   3225: 'Carrier 50 Drive: PROFINET Setpoint timeout', class No Acknowledgement, trigger "DB302_HMI_Faults_Carrier50_Faults_1" bit 8
   3226: 'Carrier 50 Power unit: Overcurrent', class No Acknowledgement, trigger "DB302_HMI_Faults_Carrier50_Faults_1" bit 9
   3227: 'Carrier 50 Power unit: DC link voltage overvoltage', class No Acknowledgement, trigger "DB302_HMI_Faults_Carrier50_Faults_1" bit 10
   3228: 'Carrier 50 Power unit: DC link voltage undervoltage', class No Acknowledgement, trigger "DB302_HMI_Faults_Carrier50_Faults_1" bit 11
   3229: 'Carrier 50 Power unit: Line phase failure in main circuit', class No Acknowledgement, trigger "DB302_HMI_Faults_Carrier50_Faults_1" bit 12
   3230: 'Carrier 50 Power unit: Phase failure motor cable', class No Acknowledgement, trigger "DB302_HMI_Faults_Carrier50_Faults_1" bit 13
   3231: 'Carrier 50 Power unit: Ground fault', class No Acknowledgement, trigger "DB302_HMI_Faults_Carrier50_Faults_1" bit 14
   3232: 'Spare_Fault_3232', class No Acknowledgement, trigger "DB302_HMI_Faults_Carrier50_Faults_1" bit 15
   3233: 'Carrier 50 Motion Off Fault', class No Acknowledgement, trigger "DB302_HMI_Faults_Carrier50_Faults_2" bit 0
   3234: 'Carrier 50 Motion On Fault', class No Acknowledgement, trigger "DB302_HMI_Faults_Carrier50_Faults_2" bit 1
   3235: 'Carrier 50 Spacing Fault', class No Acknowledgement, trigger "DB302_HMI_Faults_Carrier50_Faults_2" bit 2
   3236: 'Carrier 50 Duplicate Carrier Number Fault', class No Acknowledgement, trigger "DB302_HMI_Faults_Carrier50_Faults_2" bit 3
   3237: 'Spare_Fault_3237', class No Acknowledgement, trigger "DB302_HMI_Faults_Carrier50_Faults_2" bit 4
   3238: 'Spare_Fault_3238', class No Acknowledgement, trigger "DB302_HMI_Faults_Carrier50_Faults_2" bit 5
   3239: 'Spare_Fault_3239', class No Acknowledgement, trigger "DB302_HMI_Faults_Carrier50_Faults_2" bit 6
   3240: 'Spare_Fault_3240', class No Acknowledgement, trigger "DB302_HMI_Faults_Carrier50_Faults_2" bit 7
   3241: 'Spare_Fault_3241', class No Acknowledgement, trigger "DB302_HMI_Faults_Carrier50_Faults_2" bit 8
   3242: 'Spare_Fault_3242', class No Acknowledgement, trigger "DB302_HMI_Faults_Carrier50_Faults_2" bit 9
   3243: 'Spare_Fault_3243', class No Acknowledgement, trigger "DB302_HMI_Faults_Carrier50_Faults_2" bit 10
   3244: 'Spare_Fault_3244', class No Acknowledgement, trigger "DB302_HMI_Faults_Carrier50_Faults_2" bit 11
   3245: 'Spare_Fault_3245', class No Acknowledgement, trigger "DB302_HMI_Faults_Carrier50_Faults_2" bit 12
   3246: 'Spare_Fault_3246', class No Acknowledgement, trigger "DB302_HMI_Faults_Carrier50_Faults_2" bit 13
   3247: 'Spare_Fault_3247', class No Acknowledgement, trigger "DB302_HMI_Faults_Carrier50_Faults_2" bit 14
   3248: 'Spare_Fault_3248', class No Acknowledgement, trigger "DB302_HMI_Faults_Carrier50_Faults_2" bit 15
   3249: 'Spare_Fault_3249', class No Acknowledgement, trigger "DB302_HMI_Faults_Carrier50_Faults_3" bit 0
   3250: 'Spare_Fault_3250', class No Acknowledgement, trigger "DB302_HMI_Faults_Carrier50_Faults_3" bit 1
   3251: 'Spare_Fault_3251', class No Acknowledgement, trigger "DB302_HMI_Faults_Carrier50_Faults_3" bit 2
   3252: 'Spare_Fault_3252', class No Acknowledgement, trigger "DB302_HMI_Faults_Carrier50_Faults_3" bit 3
   3253: 'Spare_Fault_3253', class No Acknowledgement, trigger "DB302_HMI_Faults_Carrier50_Faults_3" bit 4
   3254: 'Spare_Fault_3254', class No Acknowledgement, trigger "DB302_HMI_Faults_Carrier50_Faults_3" bit 5
   3255: 'Spare_Fault_3255', class No Acknowledgement, trigger "DB302_HMI_Faults_Carrier50_Faults_3" bit 6
   3256: 'Spare_Fault_3256', class No Acknowledgement, trigger "DB302_HMI_Faults_Carrier50_Faults_3" bit 7
   3257: 'Spare_Fault_3257', class No Acknowledgement, trigger "DB302_HMI_Faults_Carrier50_Faults_3" bit 8
   3258: 'Spare_Fault_3258', class No Acknowledgement, trigger "DB302_HMI_Faults_Carrier50_Faults_3" bit 9
   3259: 'Spare_Fault_3259', class No Acknowledgement, trigger "DB302_HMI_Faults_Carrier50_Faults_3" bit 10
   3260: 'Spare_Fault_3260', class No Acknowledgement, trigger "DB302_HMI_Faults_Carrier50_Faults_3" bit 11
   3261: 'Spare_Fault_3261', class No Acknowledgement, trigger "DB302_HMI_Faults_Carrier50_Faults_3" bit 12
   3262: 'Spare_Fault_3262', class No Acknowledgement, trigger "DB302_HMI_Faults_Carrier50_Faults_3" bit 13
   3263: 'Spare_Fault_3263', class No Acknowledgement, trigger "DB302_HMI_Faults_Carrier50_Faults_3" bit 14
   3264: 'Spare_Fault_3264', class No Acknowledgement, trigger "DB302_HMI_Faults_Carrier50_Faults_3" bit 15
   3265: 'Carrier 51 Disconnect Open Power Fault DI11.0', class No Acknowledgement, trigger "DB302_HMI_Faults_Carrier51_Faults_0" bit 0
   3266: 'Carrier 51 Drive Profinet Comm Fault', class No Acknowledgement, trigger "DB302_HMI_Faults_Carrier51_Faults_0" bit 1
   3267: 'Carrier 51 Production Stop Not Reset', class No Acknowledgement, trigger "DB302_HMI_Faults_Carrier51_Faults_0" bit 2
   3268: 'Carrier 51 CB02122 Tripped', class No Acknowledgement, trigger "DB302_HMI_Faults_Carrier51_Faults_0" bit 3
   3269: 'Carrier 51 CB02123 Tripped', class No Acknowledgement, trigger "DB302_HMI_Faults_Carrier51_Faults_0" bit 4
   3270: 'Carrier 51 AUX1 CB Tripped', class No Acknowledgement, trigger "DB302_HMI_Faults_Carrier51_Faults_0" bit 5
   3271: 'Carrier 51 AUX2 CB Tripped', class No Acknowledgement, trigger "DB302_HMI_Faults_Carrier51_Faults_0" bit 6
   3272: 'Carrier 51 PLC Not Communicating', class No Acknowledgement, trigger "DB302_HMI_Faults_Carrier51_Faults_0" bit 7
   3273: 'Carrier 51 Safe Input Card Fault', class No Acknowledgement, trigger "DB302_HMI_Faults_Carrier51_Faults_0" bit 8
   3274: 'Carrier 51 Safe Output Card Fault', class No Acknowledgement, trigger "DB302_HMI_Faults_Carrier51_Faults_0" bit 9
   3275: 'Carrier 51 Standard Input Card Fault', class No Acknowledgement, trigger "DB302_HMI_Faults_Carrier51_Faults_0" bit 10
   3276: 'Carrier 51 Standard Output Card Fault', class No Acknowledgement, trigger "DB302_HMI_Faults_Carrier51_Faults_0" bit 11
   3277: 'Carrier 51 Encoder Position Fault', class No Acknowledgement, trigger "DB302_HMI_Faults_Carrier51_Faults_0" bit 12
   3278: 'Carrier 51 Encoder Internal Error', class No Acknowledgement, trigger "DB302_HMI_Faults_Carrier51_Faults_0" bit 13
   3279: 'Carrier 51 Encoder Comm Fault', class No Acknowledgement, trigger "DB302_HMI_Faults_Carrier51_Faults_0" bit 14
   3280: 'Carrier 51 HMI Comm Fault', class No Acknowledgement, trigger "DB302_HMI_Faults_Carrier51_Faults_0" bit 15
   3281: 'Carrier 51 Crash Detection Fault', class No Acknowledgement, trigger "DB302_HMI_Faults_Carrier51_Faults_1" bit 0
   3282: 'Carrier 51 Carrier Number Invalid', class No Acknowledgement, trigger "DB302_HMI_Faults_Carrier51_Faults_1" bit 1
   3283: 'Carrier 51 Drive: PROFINET configuration error', class No Acknowledgement, trigger "DB302_HMI_Faults_Carrier51_Faults_1" bit 2
   3284: 'Carrier 51 Drive: Error internal communications', class No Acknowledgement, trigger "DB302_HMI_Faults_Carrier51_Faults_1" bit 3
   3285: 'Carrier 51 Drive: Motor overtemperature', class No Acknowledgement, trigger "DB302_HMI_Faults_Carrier51_Faults_1" bit 4
   3286: 'Carrier 51 Drive: Motor overcurrent', class No Acknowledgement, trigger "DB302_HMI_Faults_Carrier51_Faults_1" bit 5
   3287: 'Carrier 51 Drive: Infeed or power unit not ready', class No Acknowledgement, trigger "DB302_HMI_Faults_Carrier51_Faults_1" bit 6
   3288: 'Carrier 51 Drive: Short-circuit/ground fault detected', class No Acknowledgement, trigger "DB302_HMI_Faults_Carrier51_Faults_1" bit 7
   3289: 'Carrier 51 Drive: PROFINET Setpoint timeout', class No Acknowledgement, trigger "DB302_HMI_Faults_Carrier51_Faults_1" bit 8
   3290: 'Carrier 51 Power unit: Overcurrent', class No Acknowledgement, trigger "DB302_HMI_Faults_Carrier51_Faults_1" bit 9
   3291: 'Carrier 51 Power unit: DC link voltage overvoltage', class No Acknowledgement, trigger "DB302_HMI_Faults_Carrier51_Faults_1" bit 10
   3292: 'Carrier 51 Power unit: DC link voltage undervoltage', class No Acknowledgement, trigger "DB302_HMI_Faults_Carrier51_Faults_1" bit 11
   3293: 'Carrier 51 Power unit: Line phase failure in main circuit', class No Acknowledgement, trigger "DB302_HMI_Faults_Carrier51_Faults_1" bit 12
   3294: 'Carrier 51 Power unit: Phase failure motor cable', class No Acknowledgement, trigger "DB302_HMI_Faults_Carrier51_Faults_1" bit 13
   3295: 'Carrier 51 Power unit: Ground fault', class No Acknowledgement, trigger "DB302_HMI_Faults_Carrier51_Faults_1" bit 14
   3296: 'Spare_Fault_3296', class No Acknowledgement, trigger "DB302_HMI_Faults_Carrier51_Faults_1" bit 15
   3297: 'Carrier 51 Motion Off Fault', class No Acknowledgement, trigger "DB302_HMI_Faults_Carrier51_Faults_2" bit 0
   3298: 'Carrier 51 Motion On Fault', class No Acknowledgement, trigger "DB302_HMI_Faults_Carrier51_Faults_2" bit 1
   3299: 'Carrier 51 Spacing Fault', class No Acknowledgement, trigger "DB302_HMI_Faults_Carrier51_Faults_2" bit 2
   3300: 'Carrier 51 Duplicate Carrier Number Fault', class No Acknowledgement, trigger "DB302_HMI_Faults_Carrier51_Faults_2" bit 3
   3301: 'Spare_Fault_3301', class No Acknowledgement, trigger "DB302_HMI_Faults_Carrier51_Faults_2" bit 4
   3302: 'Spare_Fault_3302', class No Acknowledgement, trigger "DB302_HMI_Faults_Carrier51_Faults_2" bit 5
   3303: 'Spare_Fault_3303', class No Acknowledgement, trigger "DB302_HMI_Faults_Carrier51_Faults_2" bit 6
   3304: 'Spare_Fault_3304', class No Acknowledgement, trigger "DB302_HMI_Faults_Carrier51_Faults_2" bit 7
   3305: 'Spare_Fault_3305', class No Acknowledgement, trigger "DB302_HMI_Faults_Carrier51_Faults_2" bit 8
   3306: 'Spare_Fault_3306', class No Acknowledgement, trigger "DB302_HMI_Faults_Carrier51_Faults_2" bit 9
   3307: 'Spare_Fault_3307', class No Acknowledgement, trigger "DB302_HMI_Faults_Carrier51_Faults_2" bit 10
   3308: 'Spare_Fault_3308', class No Acknowledgement, trigger "DB302_HMI_Faults_Carrier51_Faults_2" bit 11
   3309: 'Spare_Fault_3309', class No Acknowledgement, trigger "DB302_HMI_Faults_Carrier51_Faults_2" bit 12
   3310: 'Spare_Fault_3310', class No Acknowledgement, trigger "DB302_HMI_Faults_Carrier51_Faults_2" bit 13
   3311: 'Spare_Fault_3311', class No Acknowledgement, trigger "DB302_HMI_Faults_Carrier51_Faults_2" bit 14
   3312: 'Spare_Fault_3312', class No Acknowledgement, trigger "DB302_HMI_Faults_Carrier51_Faults_2" bit 15
   3313: 'Spare_Fault_3313', class No Acknowledgement, trigger "DB302_HMI_Faults_Carrier51_Faults_3" bit 0
   3314: 'Spare_Fault_3314', class No Acknowledgement, trigger "DB302_HMI_Faults_Carrier51_Faults_3" bit 1
   3315: 'Spare_Fault_3315', class No Acknowledgement, trigger "DB302_HMI_Faults_Carrier51_Faults_3" bit 2
   3316: 'Spare_Fault_3316', class No Acknowledgement, trigger "DB302_HMI_Faults_Carrier51_Faults_3" bit 3
   3317: 'Spare_Fault_3317', class No Acknowledgement, trigger "DB302_HMI_Faults_Carrier51_Faults_3" bit 4
   3318: 'Spare_Fault_3318', class No Acknowledgement, trigger "DB302_HMI_Faults_Carrier51_Faults_3" bit 5
   3319: 'Spare_Fault_3319', class No Acknowledgement, trigger "DB302_HMI_Faults_Carrier51_Faults_3" bit 6
   3320: 'Spare_Fault_3320', class No Acknowledgement, trigger "DB302_HMI_Faults_Carrier51_Faults_3" bit 7
   3321: 'Spare_Fault_3321', class No Acknowledgement, trigger "DB302_HMI_Faults_Carrier51_Faults_3" bit 8
   3322: 'Spare_Fault_3322', class No Acknowledgement, trigger "DB302_HMI_Faults_Carrier51_Faults_3" bit 9
   3323: 'Spare_Fault_3323', class No Acknowledgement, trigger "DB302_HMI_Faults_Carrier51_Faults_3" bit 10
   3324: 'Spare_Fault_3324', class No Acknowledgement, trigger "DB302_HMI_Faults_Carrier51_Faults_3" bit 11
   3325: 'Spare_Fault_3325', class No Acknowledgement, trigger "DB302_HMI_Faults_Carrier51_Faults_3" bit 12
   3326: 'Spare_Fault_3326', class No Acknowledgement, trigger "DB302_HMI_Faults_Carrier51_Faults_3" bit 13
   3327: 'Spare_Fault_3327', class No Acknowledgement, trigger "DB302_HMI_Faults_Carrier51_Faults_3" bit 14
   3328: 'Spare_Fault_3328', class No Acknowledgement, trigger "DB302_HMI_Faults_Carrier51_Faults_3" bit 15
   3329: 'Carrier 52 Disconnect Open Power Fault DI11.0', class No Acknowledgement, trigger "DB302_HMI_Faults_Carrier52_Faults_0" bit 0
   3330: 'Carrier 52 Drive Profinet Comm Fault', class No Acknowledgement, trigger "DB302_HMI_Faults_Carrier52_Faults_0" bit 1
   3331: 'Carrier 52 Production Stop Not Reset', class No Acknowledgement, trigger "DB302_HMI_Faults_Carrier52_Faults_0" bit 2
   3332: 'Carrier 52 CB02122 Tripped', class No Acknowledgement, trigger "DB302_HMI_Faults_Carrier52_Faults_0" bit 3
   3333: 'Carrier 52 CB02123 Tripped', class No Acknowledgement, trigger "DB302_HMI_Faults_Carrier52_Faults_0" bit 4
   3334: 'Carrier 52 AUX1 CB Tripped', class No Acknowledgement, trigger "DB302_HMI_Faults_Carrier52_Faults_0" bit 5
   3335: 'Carrier 52 AUX2 CB Tripped', class No Acknowledgement, trigger "DB302_HMI_Faults_Carrier52_Faults_0" bit 6
   3336: 'Carrier 52 PLC Not Communicating', class No Acknowledgement, trigger "DB302_HMI_Faults_Carrier52_Faults_0" bit 7
   3337: 'Carrier 52 Safe Input Card Fault', class No Acknowledgement, trigger "DB302_HMI_Faults_Carrier52_Faults_0" bit 8
   3338: 'Carrier 52 Safe Output Card Fault', class No Acknowledgement, trigger "DB302_HMI_Faults_Carrier52_Faults_0" bit 9
   3339: 'Carrier 52 Standard Input Card Fault', class No Acknowledgement, trigger "DB302_HMI_Faults_Carrier52_Faults_0" bit 10
   3340: 'Carrier 52 Standard Output Card Fault', class No Acknowledgement, trigger "DB302_HMI_Faults_Carrier52_Faults_0" bit 11
   3341: 'Carrier 52 Encoder Position Fault', class No Acknowledgement, trigger "DB302_HMI_Faults_Carrier52_Faults_0" bit 12
   3342: 'Carrier 52 Encoder Internal Error', class No Acknowledgement, trigger "DB302_HMI_Faults_Carrier52_Faults_0" bit 13
   3343: 'Carrier 52 Encoder Comm Fault', class No Acknowledgement, trigger "DB302_HMI_Faults_Carrier52_Faults_0" bit 14
   3344: 'Carrier 52 HMI Comm Fault', class No Acknowledgement, trigger "DB302_HMI_Faults_Carrier52_Faults_0" bit 15
   3345: 'Carrier 52 Crash Detection Fault', class No Acknowledgement, trigger "DB302_HMI_Faults_Carrier52_Faults_1" bit 0
   3346: 'Carrier 52 Carrier Number Invalid', class No Acknowledgement, trigger "DB302_HMI_Faults_Carrier52_Faults_1" bit 1
   3347: 'Carrier 52 Drive: PROFINET configuration error', class No Acknowledgement, trigger "DB302_HMI_Faults_Carrier52_Faults_1" bit 2
   3348: 'Carrier 52 Drive: Error internal communications', class No Acknowledgement, trigger "DB302_HMI_Faults_Carrier52_Faults_1" bit 3
   3349: 'Carrier 52 Drive: Motor overtemperature', class No Acknowledgement, trigger "DB302_HMI_Faults_Carrier52_Faults_1" bit 4
   3350: 'Carrier 52 Drive: Motor overcurrent', class No Acknowledgement, trigger "DB302_HMI_Faults_Carrier52_Faults_1" bit 5
   3351: 'Carrier 52 Drive: Infeed or power unit not ready', class No Acknowledgement, trigger "DB302_HMI_Faults_Carrier52_Faults_1" bit 6
   3352: 'Carrier 52 Drive: Short-circuit/ground fault detected', class No Acknowledgement, trigger "DB302_HMI_Faults_Carrier52_Faults_1" bit 7
   3353: 'Carrier 52 Drive: PROFINET Setpoint timeout', class No Acknowledgement, trigger "DB302_HMI_Faults_Carrier52_Faults_1" bit 8
   3354: 'Carrier 52 Power unit: Overcurrent', class No Acknowledgement, trigger "DB302_HMI_Faults_Carrier52_Faults_1" bit 9
   3355: 'Carrier 52 Power unit: DC link voltage overvoltage', class No Acknowledgement, trigger "DB302_HMI_Faults_Carrier52_Faults_1" bit 10
   3356: 'Carrier 52 Power unit: DC link voltage undervoltage', class No Acknowledgement, trigger "DB302_HMI_Faults_Carrier52_Faults_1" bit 11
   3357: 'Carrier 52 Power unit: Line phase failure in main circuit', class No Acknowledgement, trigger "DB302_HMI_Faults_Carrier52_Faults_1" bit 12
   3358: 'Carrier 52 Power unit: Phase failure motor cable', class No Acknowledgement, trigger "DB302_HMI_Faults_Carrier52_Faults_1" bit 13
   3359: 'Carrier 52 Power unit: Ground fault', class No Acknowledgement, trigger "DB302_HMI_Faults_Carrier52_Faults_1" bit 14
   3360: 'Spare_Fault_3360', class No Acknowledgement, trigger "DB302_HMI_Faults_Carrier52_Faults_1" bit 15
   3361: 'Carrier 52 Motion Off Fault', class No Acknowledgement, trigger "DB302_HMI_Faults_Carrier52_Faults_2" bit 0
   3362: 'Carrier 52 Motion On Fault', class No Acknowledgement, trigger "DB302_HMI_Faults_Carrier52_Faults_2" bit 1
   3363: 'Carrier 52 Spacing Fault', class No Acknowledgement, trigger "DB302_HMI_Faults_Carrier52_Faults_2" bit 2
   3364: 'Carrier 52 Duplicate Carrier Number Fault', class No Acknowledgement, trigger "DB302_HMI_Faults_Carrier52_Faults_2" bit 3
   3365: 'Spare_Fault_3365', class No Acknowledgement, trigger "DB302_HMI_Faults_Carrier52_Faults_2" bit 4
   3366: 'Spare_Fault_3366', class No Acknowledgement, trigger "DB302_HMI_Faults_Carrier52_Faults_2" bit 5
   3367: 'Spare_Fault_3367', class No Acknowledgement, trigger "DB302_HMI_Faults_Carrier52_Faults_2" bit 6
   3368: 'Spare_Fault_3368', class No Acknowledgement, trigger "DB302_HMI_Faults_Carrier52_Faults_2" bit 7
   3369: 'Spare_Fault_3369', class No Acknowledgement, trigger "DB302_HMI_Faults_Carrier52_Faults_2" bit 8
   3370: 'Spare_Fault_3370', class No Acknowledgement, trigger "DB302_HMI_Faults_Carrier52_Faults_2" bit 9
   3371: 'Spare_Fault_3371', class No Acknowledgement, trigger "DB302_HMI_Faults_Carrier52_Faults_2" bit 10
   3372: 'Spare_Fault_3372', class No Acknowledgement, trigger "DB302_HMI_Faults_Carrier52_Faults_2" bit 11
   3373: 'Spare_Fault_3373', class No Acknowledgement, trigger "DB302_HMI_Faults_Carrier52_Faults_2" bit 12
   3374: 'Spare_Fault_3374', class No Acknowledgement, trigger "DB302_HMI_Faults_Carrier52_Faults_2" bit 13
   3375: 'Spare_Fault_3375', class No Acknowledgement, trigger "DB302_HMI_Faults_Carrier52_Faults_2" bit 14
   3376: 'Spare_Fault_3376', class No Acknowledgement, trigger "DB302_HMI_Faults_Carrier52_Faults_2" bit 15
   3377: 'Spare_Fault_3377', class No Acknowledgement, trigger "DB302_HMI_Faults_Carrier52_Faults_3" bit 0
   3378: 'Spare_Fault_3378', class No Acknowledgement, trigger "DB302_HMI_Faults_Carrier52_Faults_3" bit 1
   3379: 'Spare_Fault_3379', class No Acknowledgement, trigger "DB302_HMI_Faults_Carrier52_Faults_3" bit 2
   3380: 'Spare_Fault_3380', class No Acknowledgement, trigger "DB302_HMI_Faults_Carrier52_Faults_3" bit 3
   3381: 'Spare_Fault_3381', class No Acknowledgement, trigger "DB302_HMI_Faults_Carrier52_Faults_3" bit 4
   3382: 'Spare_Fault_3382', class No Acknowledgement, trigger "DB302_HMI_Faults_Carrier52_Faults_3" bit 5
   3383: 'Spare_Fault_3383', class No Acknowledgement, trigger "DB302_HMI_Faults_Carrier52_Faults_3" bit 6
   3384: 'Spare_Fault_3384', class No Acknowledgement, trigger "DB302_HMI_Faults_Carrier52_Faults_3" bit 7
   3385: 'Spare_Fault_3385', class No Acknowledgement, trigger "DB302_HMI_Faults_Carrier52_Faults_3" bit 8
   3386: 'Spare_Fault_3386', class No Acknowledgement, trigger "DB302_HMI_Faults_Carrier52_Faults_3" bit 9
   3387: 'Spare_Fault_3387', class No Acknowledgement, trigger "DB302_HMI_Faults_Carrier52_Faults_3" bit 10
   3388: 'Spare_Fault_3388', class No Acknowledgement, trigger "DB302_HMI_Faults_Carrier52_Faults_3" bit 11
   3389: 'Spare_Fault_3389', class No Acknowledgement, trigger "DB302_HMI_Faults_Carrier52_Faults_3" bit 12
   3390: 'Spare_Fault_3390', class No Acknowledgement, trigger "DB302_HMI_Faults_Carrier52_Faults_3" bit 13
   3391: 'Spare_Fault_3391', class No Acknowledgement, trigger "DB302_HMI_Faults_Carrier52_Faults_3" bit 14
   3392: 'Spare_Fault_3392', class No Acknowledgement, trigger "DB302_HMI_Faults_Carrier52_Faults_3" bit 15
   3393: 'Carrier 53 Disconnect Open Power Fault DI11.0', class No Acknowledgement, trigger "DB302_HMI_Faults_Carrier53_Faults_0" bit 0
   3394: 'Carrier 53 Drive Profinet Comm Fault', class No Acknowledgement, trigger "DB302_HMI_Faults_Carrier53_Faults_0" bit 1
   3395: 'Carrier 53 Production Stop Not Reset', class No Acknowledgement, trigger "DB302_HMI_Faults_Carrier53_Faults_0" bit 2
   3396: 'Carrier 53 CB02122 Tripped', class No Acknowledgement, trigger "DB302_HMI_Faults_Carrier53_Faults_0" bit 3
   3397: 'Carrier 53 CB02123 Tripped', class No Acknowledgement, trigger "DB302_HMI_Faults_Carrier53_Faults_0" bit 4
   3398: 'Carrier 53 AUX1 CB Tripped', class No Acknowledgement, trigger "DB302_HMI_Faults_Carrier53_Faults_0" bit 5
   3399: 'Carrier 53 AUX2 CB Tripped', class No Acknowledgement, trigger "DB302_HMI_Faults_Carrier53_Faults_0" bit 6
   3400: 'Carrier 53 PLC Not Communicating', class No Acknowledgement, trigger "DB302_HMI_Faults_Carrier53_Faults_0" bit 7
   3401: 'Carrier 53 Safe Input Card Fault', class No Acknowledgement, trigger "DB302_HMI_Faults_Carrier53_Faults_0" bit 8
   3402: 'Carrier 53 Safe Output Card Fault', class No Acknowledgement, trigger "DB302_HMI_Faults_Carrier53_Faults_0" bit 9
   3403: 'Carrier 53 Standard Input Card Fault', class No Acknowledgement, trigger "DB302_HMI_Faults_Carrier53_Faults_0" bit 10
   3404: 'Carrier 53 Standard Output Card Fault', class No Acknowledgement, trigger "DB302_HMI_Faults_Carrier53_Faults_0" bit 11
   3405: 'Carrier 53 Encoder Position Fault', class No Acknowledgement, trigger "DB302_HMI_Faults_Carrier53_Faults_0" bit 12
   3406: 'Carrier 53 Encoder Internal Error', class No Acknowledgement, trigger "DB302_HMI_Faults_Carrier53_Faults_0" bit 13
   3407: 'Carrier 53 Encoder Comm Fault', class No Acknowledgement, trigger "DB302_HMI_Faults_Carrier53_Faults_0" bit 14
   3408: 'Carrier 53 HMI Comm Fault', class No Acknowledgement, trigger "DB302_HMI_Faults_Carrier53_Faults_0" bit 15
   3409: 'Carrier 53 Crash Detection Fault', class No Acknowledgement, trigger "DB302_HMI_Faults_Carrier53_Faults_1" bit 0
   3410: 'Carrier 53 Carrier Number Invalid', class No Acknowledgement, trigger "DB302_HMI_Faults_Carrier53_Faults_1" bit 1
   3411: 'Carrier 53 Drive: PROFINET configuration error', class No Acknowledgement, trigger "DB302_HMI_Faults_Carrier53_Faults_1" bit 2
   3412: 'Carrier 53 Drive: Error internal communications', class No Acknowledgement, trigger "DB302_HMI_Faults_Carrier53_Faults_1" bit 3
   3413: 'Carrier 53 Drive: Motor overtemperature', class No Acknowledgement, trigger "DB302_HMI_Faults_Carrier53_Faults_1" bit 4
   3414: 'Carrier 53 Drive: Motor overcurrent', class No Acknowledgement, trigger "DB302_HMI_Faults_Carrier53_Faults_1" bit 5
   3415: 'Carrier 53 Drive: Infeed or power unit not ready', class No Acknowledgement, trigger "DB302_HMI_Faults_Carrier53_Faults_1" bit 6
   3416: 'Carrier 53 Drive: Short-circuit/ground fault detected', class No Acknowledgement, trigger "DB302_HMI_Faults_Carrier53_Faults_1" bit 7
   3417: 'Carrier 53 Drive: PROFINET Setpoint timeout', class No Acknowledgement, trigger "DB302_HMI_Faults_Carrier53_Faults_1" bit 8
   3418: 'Carrier 53 Power unit: Overcurrent', class No Acknowledgement, trigger "DB302_HMI_Faults_Carrier53_Faults_1" bit 9
   3419: 'Carrier 53 Power unit: DC link voltage overvoltage', class No Acknowledgement, trigger "DB302_HMI_Faults_Carrier53_Faults_1" bit 10
   3420: 'Carrier 53 Power unit: DC link voltage undervoltage', class No Acknowledgement, trigger "DB302_HMI_Faults_Carrier53_Faults_1" bit 11
   3421: 'Carrier 53 Power unit: Line phase failure in main circuit', class No Acknowledgement, trigger "DB302_HMI_Faults_Carrier53_Faults_1" bit 12
   3422: 'Carrier 53 Power unit: Phase failure motor cable', class No Acknowledgement, trigger "DB302_HMI_Faults_Carrier53_Faults_1" bit 13
   3423: 'Carrier 53 Power unit: Ground fault', class No Acknowledgement, trigger "DB302_HMI_Faults_Carrier53_Faults_1" bit 14
   3424: 'Spare_Fault_3424', class No Acknowledgement, trigger "DB302_HMI_Faults_Carrier53_Faults_1" bit 15
   3425: 'Carrier 53 Motion Off Fault', class No Acknowledgement, trigger "DB302_HMI_Faults_Carrier53_Faults_2" bit 0
   3426: 'Carrier 53 Motion On Fault', class No Acknowledgement, trigger "DB302_HMI_Faults_Carrier53_Faults_2" bit 1
   3427: 'Carrier 53 Spacing Fault', class No Acknowledgement, trigger "DB302_HMI_Faults_Carrier53_Faults_2" bit 2
   3428: 'Carrier 53 Duplicate Carrier Number Fault', class No Acknowledgement, trigger "DB302_HMI_Faults_Carrier53_Faults_2" bit 3
   3429: 'Spare_Fault_3429', class No Acknowledgement, trigger "DB302_HMI_Faults_Carrier53_Faults_2" bit 4
   3430: 'Spare_Fault_3430', class No Acknowledgement, trigger "DB302_HMI_Faults_Carrier53_Faults_2" bit 5
   3431: 'Spare_Fault_3431', class No Acknowledgement, trigger "DB302_HMI_Faults_Carrier53_Faults_2" bit 6
   3432: 'Spare_Fault_3432', class No Acknowledgement, trigger "DB302_HMI_Faults_Carrier53_Faults_2" bit 7
   3433: 'Spare_Fault_3433', class No Acknowledgement, trigger "DB302_HMI_Faults_Carrier53_Faults_2" bit 8
   3434: 'Spare_Fault_3434', class No Acknowledgement, trigger "DB302_HMI_Faults_Carrier53_Faults_2" bit 9
   3435: 'Spare_Fault_3435', class No Acknowledgement, trigger "DB302_HMI_Faults_Carrier53_Faults_2" bit 10
   3436: 'Spare_Fault_3436', class No Acknowledgement, trigger "DB302_HMI_Faults_Carrier53_Faults_2" bit 11
   3437: 'Spare_Fault_3437', class No Acknowledgement, trigger "DB302_HMI_Faults_Carrier53_Faults_2" bit 12
   3438: 'Spare_Fault_3438', class No Acknowledgement, trigger "DB302_HMI_Faults_Carrier53_Faults_2" bit 13
   3439: 'Spare_Fault_3439', class No Acknowledgement, trigger "DB302_HMI_Faults_Carrier53_Faults_2" bit 14
   3440: 'Spare_Fault_3440', class No Acknowledgement, trigger "DB302_HMI_Faults_Carrier53_Faults_2" bit 15
   3441: 'Spare_Fault_3441', class No Acknowledgement, trigger "DB302_HMI_Faults_Carrier53_Faults_3" bit 0
   3442: 'Spare_Fault_3442', class No Acknowledgement, trigger "DB302_HMI_Faults_Carrier53_Faults_3" bit 1
   3443: 'Spare_Fault_3443', class No Acknowledgement, trigger "DB302_HMI_Faults_Carrier53_Faults_3" bit 2
   3444: 'Spare_Fault_3444', class No Acknowledgement, trigger "DB302_HMI_Faults_Carrier53_Faults_3" bit 3
   3445: 'Spare_Fault_3445', class No Acknowledgement, trigger "DB302_HMI_Faults_Carrier53_Faults_3" bit 4
   3446: 'Spare_Fault_3446', class No Acknowledgement, trigger "DB302_HMI_Faults_Carrier53_Faults_3" bit 5
   3447: 'Spare_Fault_3447', class No Acknowledgement, trigger "DB302_HMI_Faults_Carrier53_Faults_3" bit 6
   3448: 'Spare_Fault_3448', class No Acknowledgement, trigger "DB302_HMI_Faults_Carrier53_Faults_3" bit 7
   3449: 'Spare_Fault_3449', class No Acknowledgement, trigger "DB302_HMI_Faults_Carrier53_Faults_3" bit 8
   3450: 'Spare_Fault_3450', class No Acknowledgement, trigger "DB302_HMI_Faults_Carrier53_Faults_3" bit 9
   3451: 'Spare_Fault_3451', class No Acknowledgement, trigger "DB302_HMI_Faults_Carrier53_Faults_3" bit 10
   3452: 'Spare_Fault_3452', class No Acknowledgement, trigger "DB302_HMI_Faults_Carrier53_Faults_3" bit 11
   3453: 'Spare_Fault_3453', class No Acknowledgement, trigger "DB302_HMI_Faults_Carrier53_Faults_3" bit 12
   3454: 'Spare_Fault_3454', class No Acknowledgement, trigger "DB302_HMI_Faults_Carrier53_Faults_3" bit 13
   3455: 'Spare_Fault_3455', class No Acknowledgement, trigger "DB302_HMI_Faults_Carrier53_Faults_3" bit 14
   3456: 'Spare_Fault_3456', class No Acknowledgement, trigger "DB302_HMI_Faults_Carrier53_Faults_3" bit 15
   3457: 'Carrier 54 Disconnect Open Power Fault DI11.0', class No Acknowledgement, trigger "DB302_HMI_Faults_Carrier54_Faults_0" bit 0
   3458: 'Carrier 54 Drive Profinet Comm Fault', class No Acknowledgement, trigger "DB302_HMI_Faults_Carrier54_Faults_0" bit 1
   3459: 'Carrier 54 Production Stop Not Reset', class No Acknowledgement, trigger "DB302_HMI_Faults_Carrier54_Faults_0" bit 2
   3460: 'Carrier 54 CB02122 Tripped', class No Acknowledgement, trigger "DB302_HMI_Faults_Carrier54_Faults_0" bit 3
   3461: 'Carrier 54 CB02123 Tripped', class No Acknowledgement, trigger "DB302_HMI_Faults_Carrier54_Faults_0" bit 4
   3462: 'Carrier 54 AUX1 CB Tripped', class No Acknowledgement, trigger "DB302_HMI_Faults_Carrier54_Faults_0" bit 5
   3463: 'Carrier 54 AUX2 CB Tripped', class No Acknowledgement, trigger "DB302_HMI_Faults_Carrier54_Faults_0" bit 6
   3464: 'Carrier 54 PLC Not Communicating', class No Acknowledgement, trigger "DB302_HMI_Faults_Carrier54_Faults_0" bit 7
   3465: 'Carrier 54 Safe Input Card Fault', class No Acknowledgement, trigger "DB302_HMI_Faults_Carrier54_Faults_0" bit 8
   3466: 'Carrier 54 Safe Output Card Fault', class No Acknowledgement, trigger "DB302_HMI_Faults_Carrier54_Faults_0" bit 9
   3467: 'Carrier 54 Standard Input Card Fault', class No Acknowledgement, trigger "DB302_HMI_Faults_Carrier54_Faults_0" bit 10
   3468: 'Carrier 54 Standard Output Card Fault', class No Acknowledgement, trigger "DB302_HMI_Faults_Carrier54_Faults_0" bit 11
   3469: 'Carrier 54 Encoder Position Fault', class No Acknowledgement, trigger "DB302_HMI_Faults_Carrier54_Faults_0" bit 12
   3470: 'Carrier 54 Encoder Internal Error', class No Acknowledgement, trigger "DB302_HMI_Faults_Carrier54_Faults_0" bit 13
   3471: 'Carrier 54 Encoder Comm Fault', class No Acknowledgement, trigger "DB302_HMI_Faults_Carrier54_Faults_0" bit 14
   3472: 'Carrier 54 HMI Comm Fault', class No Acknowledgement, trigger "DB302_HMI_Faults_Carrier54_Faults_0" bit 15
   3473: 'Carrier 54 Crash Detection Fault', class No Acknowledgement, trigger "DB302_HMI_Faults_Carrier54_Faults_1" bit 0
   3474: 'Carrier 54 Carrier Number Invalid', class No Acknowledgement, trigger "DB302_HMI_Faults_Carrier54_Faults_1" bit 1
   3475: 'Carrier 54 Drive: PROFINET configuration error', class No Acknowledgement, trigger "DB302_HMI_Faults_Carrier54_Faults_1" bit 2
   3476: 'Carrier 54 Drive: Error internal communications', class No Acknowledgement, trigger "DB302_HMI_Faults_Carrier54_Faults_1" bit 3
   3477: 'Carrier 54 Drive: Motor overtemperature', class No Acknowledgement, trigger "DB302_HMI_Faults_Carrier54_Faults_1" bit 4
   3478: 'Carrier 54 Drive: Motor overcurrent', class No Acknowledgement, trigger "DB302_HMI_Faults_Carrier54_Faults_1" bit 5
   3479: 'Carrier 54 Drive: Infeed or power unit not ready', class No Acknowledgement, trigger "DB302_HMI_Faults_Carrier54_Faults_1" bit 6
   3480: 'Carrier 54 Drive: Short-circuit/ground fault detected', class No Acknowledgement, trigger "DB302_HMI_Faults_Carrier54_Faults_1" bit 7
   3481: 'Carrier 54 Drive: PROFINET Setpoint timeout', class No Acknowledgement, trigger "DB302_HMI_Faults_Carrier54_Faults_1" bit 8
   3482: 'Carrier 54 Power unit: Overcurrent', class No Acknowledgement, trigger "DB302_HMI_Faults_Carrier54_Faults_1" bit 9
   3483: 'Carrier 54 Power unit: DC link voltage overvoltage', class No Acknowledgement, trigger "DB302_HMI_Faults_Carrier54_Faults_1" bit 10
   3484: 'Carrier 54 Power unit: DC link voltage undervoltage', class No Acknowledgement, trigger "DB302_HMI_Faults_Carrier54_Faults_1" bit 11
   3485: 'Carrier 54 Power unit: Line phase failure in main circuit', class No Acknowledgement, trigger "DB302_HMI_Faults_Carrier54_Faults_1" bit 12
   3486: 'Carrier 54 Power unit: Phase failure motor cable', class No Acknowledgement, trigger "DB302_HMI_Faults_Carrier54_Faults_1" bit 13
   3487: 'Carrier 54 Power unit: Ground fault', class No Acknowledgement, trigger "DB302_HMI_Faults_Carrier54_Faults_1" bit 14
   3488: 'Spare_Fault_3488', class No Acknowledgement, trigger "DB302_HMI_Faults_Carrier54_Faults_1" bit 15
   3489: 'Carrier 54 Motion Off Fault', class No Acknowledgement, trigger "DB302_HMI_Faults_Carrier54_Faults_2" bit 0
   3490: 'Carrier 54 Motion On Fault', class No Acknowledgement, trigger "DB302_HMI_Faults_Carrier54_Faults_2" bit 1
   3491: 'Carrier 54 Spacing Fault', class No Acknowledgement, trigger "DB302_HMI_Faults_Carrier54_Faults_2" bit 2
   3492: 'Carrier 54 Duplicate Carrier Number Fault', class No Acknowledgement, trigger "DB302_HMI_Faults_Carrier54_Faults_2" bit 3
   3493: 'Spare_Fault_3493', class No Acknowledgement, trigger "DB302_HMI_Faults_Carrier54_Faults_2" bit 4
   3494: 'Spare_Fault_3494', class No Acknowledgement, trigger "DB302_HMI_Faults_Carrier54_Faults_2" bit 5
   3495: 'Spare_Fault_3495', class No Acknowledgement, trigger "DB302_HMI_Faults_Carrier54_Faults_2" bit 6
   3496: 'Spare_Fault_3496', class No Acknowledgement, trigger "DB302_HMI_Faults_Carrier54_Faults_2" bit 7
   3497: 'Spare_Fault_3497', class No Acknowledgement, trigger "DB302_HMI_Faults_Carrier54_Faults_2" bit 8
   3498: 'Spare_Fault_3498', class No Acknowledgement, trigger "DB302_HMI_Faults_Carrier54_Faults_2" bit 9
   3499: 'Spare_Fault_3499', class No Acknowledgement, trigger "DB302_HMI_Faults_Carrier54_Faults_2" bit 10
   3500: 'Spare_Fault_3500', class No Acknowledgement, trigger "DB302_HMI_Faults_Carrier54_Faults_2" bit 11
   3501: 'Spare_Fault_3501', class No Acknowledgement, trigger "DB302_HMI_Faults_Carrier54_Faults_2" bit 12
   3502: 'Spare_Fault_3502', class No Acknowledgement, trigger "DB302_HMI_Faults_Carrier54_Faults_2" bit 13
   3503: 'Spare_Fault_3503', class No Acknowledgement, trigger "DB302_HMI_Faults_Carrier54_Faults_2" bit 14
   3504: 'Spare_Fault_3504', class No Acknowledgement, trigger "DB302_HMI_Faults_Carrier54_Faults_2" bit 15
   3505: 'Spare_Fault_3505', class No Acknowledgement, trigger "DB302_HMI_Faults_Carrier54_Faults_3" bit 0
   3506: 'Spare_Fault_3506', class No Acknowledgement, trigger "DB302_HMI_Faults_Carrier54_Faults_3" bit 1
   3507: 'Spare_Fault_3507', class No Acknowledgement, trigger "DB302_HMI_Faults_Carrier54_Faults_3" bit 2
   3508: 'Spare_Fault_3508', class No Acknowledgement, trigger "DB302_HMI_Faults_Carrier54_Faults_3" bit 3
   3509: 'Spare_Fault_3509', class No Acknowledgement, trigger "DB302_HMI_Faults_Carrier54_Faults_3" bit 4
   3510: 'Spare_Fault_3510', class No Acknowledgement, trigger "DB302_HMI_Faults_Carrier54_Faults_3" bit 5
   3511: 'Spare_Fault_3511', class No Acknowledgement, trigger "DB302_HMI_Faults_Carrier54_Faults_3" bit 6
   3512: 'Spare_Fault_3512', class No Acknowledgement, trigger "DB302_HMI_Faults_Carrier54_Faults_3" bit 7
   3513: 'Spare_Fault_3513', class No Acknowledgement, trigger "DB302_HMI_Faults_Carrier54_Faults_3" bit 8
   3514: 'Spare_Fault_3514', class No Acknowledgement, trigger "DB302_HMI_Faults_Carrier54_Faults_3" bit 9
   3515: 'Spare_Fault_3515', class No Acknowledgement, trigger "DB302_HMI_Faults_Carrier54_Faults_3" bit 10
   3516: 'Spare_Fault_3516', class No Acknowledgement, trigger "DB302_HMI_Faults_Carrier54_Faults_3" bit 11
   3517: 'Spare_Fault_3517', class No Acknowledgement, trigger "DB302_HMI_Faults_Carrier54_Faults_3" bit 12
   3518: 'Spare_Fault_3518', class No Acknowledgement, trigger "DB302_HMI_Faults_Carrier54_Faults_3" bit 13
   3519: 'Spare_Fault_3519', class No Acknowledgement, trigger "DB302_HMI_Faults_Carrier54_Faults_3" bit 14
   3520: 'Spare_Fault_3520', class No Acknowledgement, trigger "DB302_HMI_Faults_Carrier54_Faults_3" bit 15
   3521: 'Carrier 55 Disconnect Open Power Fault DI11.0', class No Acknowledgement, trigger "DB302_HMI_Faults_Carrier55_Faults_0" bit 0
   3522: 'Carrier 55 Drive Profinet Comm Fault', class No Acknowledgement, trigger "DB302_HMI_Faults_Carrier55_Faults_0" bit 1
   3523: 'Carrier 55 Production Stop Not Reset', class No Acknowledgement, trigger "DB302_HMI_Faults_Carrier55_Faults_0" bit 2
   3524: 'Carrier 55 CB02122 Tripped', class No Acknowledgement, trigger "DB302_HMI_Faults_Carrier55_Faults_0" bit 3
   3525: 'Carrier 55 CB02123 Tripped', class No Acknowledgement, trigger "DB302_HMI_Faults_Carrier55_Faults_0" bit 4
   3526: 'Carrier 55 AUX1 CB Tripped', class No Acknowledgement, trigger "DB302_HMI_Faults_Carrier55_Faults_0" bit 5
   3527: 'Carrier 55 AUX2 CB Tripped', class No Acknowledgement, trigger "DB302_HMI_Faults_Carrier55_Faults_0" bit 6
   3528: 'Carrier 55 PLC Not Communicating', class No Acknowledgement, trigger "DB302_HMI_Faults_Carrier55_Faults_0" bit 7
   3529: 'Carrier 55 Safe Input Card Fault', class No Acknowledgement, trigger "DB302_HMI_Faults_Carrier55_Faults_0" bit 8
   3530: 'Carrier 55 Safe Output Card Fault', class No Acknowledgement, trigger "DB302_HMI_Faults_Carrier55_Faults_0" bit 9
   3531: 'Carrier 55 Standard Input Card Fault', class No Acknowledgement, trigger "DB302_HMI_Faults_Carrier55_Faults_0" bit 10
   3532: 'Carrier 55 Standard Output Card Fault', class No Acknowledgement, trigger "DB302_HMI_Faults_Carrier55_Faults_0" bit 11
   3533: 'Carrier 55 Encoder Position Fault', class No Acknowledgement, trigger "DB302_HMI_Faults_Carrier55_Faults_0" bit 12
   3534: 'Carrier 55 Encoder Internal Error', class No Acknowledgement, trigger "DB302_HMI_Faults_Carrier55_Faults_0" bit 13
   3535: 'Carrier 55 Encoder Comm Fault', class No Acknowledgement, trigger "DB302_HMI_Faults_Carrier55_Faults_0" bit 14
   3536: 'Carrier 55 HMI Comm Fault', class No Acknowledgement, trigger "DB302_HMI_Faults_Carrier55_Faults_0" bit 15
   3537: 'Carrier 55 Crash Detection Fault', class No Acknowledgement, trigger "DB302_HMI_Faults_Carrier55_Faults_1" bit 0
   3538: 'Carrier 55 Carrier Number Invalid', class No Acknowledgement, trigger "DB302_HMI_Faults_Carrier55_Faults_1" bit 1
   3539: 'Carrier 55 Drive: PROFINET configuration error', class No Acknowledgement, trigger "DB302_HMI_Faults_Carrier55_Faults_1" bit 2
   3540: 'Carrier 55 Drive: Error internal communications', class No Acknowledgement, trigger "DB302_HMI_Faults_Carrier55_Faults_1" bit 3
   3541: 'Carrier 55 Drive: Motor overtemperature', class No Acknowledgement, trigger "DB302_HMI_Faults_Carrier55_Faults_1" bit 4
   3542: 'Carrier 55 Drive: Motor overcurrent', class No Acknowledgement, trigger "DB302_HMI_Faults_Carrier55_Faults_1" bit 5
   3543: 'Carrier 55 Drive: Infeed or power unit not ready', class No Acknowledgement, trigger "DB302_HMI_Faults_Carrier55_Faults_1" bit 6
   3544: 'Carrier 55 Drive: Short-circuit/ground fault detected', class No Acknowledgement, trigger "DB302_HMI_Faults_Carrier55_Faults_1" bit 7
   3545: 'Carrier 55 Drive: PROFINET Setpoint timeout', class No Acknowledgement, trigger "DB302_HMI_Faults_Carrier55_Faults_1" bit 8
   3546: 'Carrier 55 Power unit: Overcurrent', class No Acknowledgement, trigger "DB302_HMI_Faults_Carrier55_Faults_1" bit 9
   3547: 'Carrier 55 Power unit: DC link voltage overvoltage', class No Acknowledgement, trigger "DB302_HMI_Faults_Carrier55_Faults_1" bit 10
   3548: 'Carrier 55 Power unit: DC link voltage undervoltage', class No Acknowledgement, trigger "DB302_HMI_Faults_Carrier55_Faults_1" bit 11
   3549: 'Carrier 55 Power unit: Line phase failure in main circuit', class No Acknowledgement, trigger "DB302_HMI_Faults_Carrier55_Faults_1" bit 12
   3550: 'Carrier 55 Power unit: Phase failure motor cable', class No Acknowledgement, trigger "DB302_HMI_Faults_Carrier55_Faults_1" bit 13
   3551: 'Carrier 55 Power unit: Ground fault', class No Acknowledgement, trigger "DB302_HMI_Faults_Carrier55_Faults_1" bit 14
   3552: 'Spare_Fault_3552', class No Acknowledgement, trigger "DB302_HMI_Faults_Carrier55_Faults_1" bit 15
   3553: 'Carrier 55 Motion Off Fault', class No Acknowledgement, trigger "DB302_HMI_Faults_Carrier55_Faults_2" bit 0
   3554: 'Carrier 55 Motion On Fault', class No Acknowledgement, trigger "DB302_HMI_Faults_Carrier55_Faults_2" bit 1
   3555: 'Carrier 55 Spacing Fault', class No Acknowledgement, trigger "DB302_HMI_Faults_Carrier55_Faults_2" bit 2
   3556: 'Carrier 55 Duplicate Carrier Number Fault', class No Acknowledgement, trigger "DB302_HMI_Faults_Carrier55_Faults_2" bit 3
   3557: 'Spare_Fault_3557', class No Acknowledgement, trigger "DB302_HMI_Faults_Carrier55_Faults_2" bit 4
   3558: 'Spare_Fault_3558', class No Acknowledgement, trigger "DB302_HMI_Faults_Carrier55_Faults_2" bit 5
   3559: 'Spare_Fault_3559', class No Acknowledgement, trigger "DB302_HMI_Faults_Carrier55_Faults_2" bit 6
   3560: 'Spare_Fault_3560', class No Acknowledgement, trigger "DB302_HMI_Faults_Carrier55_Faults_2" bit 7
   3561: 'Spare_Fault_3561', class No Acknowledgement, trigger "DB302_HMI_Faults_Carrier55_Faults_2" bit 8
   3562: 'Spare_Fault_3562', class No Acknowledgement, trigger "DB302_HMI_Faults_Carrier55_Faults_2" bit 9
   3563: 'Spare_Fault_3563', class No Acknowledgement, trigger "DB302_HMI_Faults_Carrier55_Faults_2" bit 10
   3564: 'Spare_Fault_3564', class No Acknowledgement, trigger "DB302_HMI_Faults_Carrier55_Faults_2" bit 11
   3565: 'Spare_Fault_3565', class No Acknowledgement, trigger "DB302_HMI_Faults_Carrier55_Faults_2" bit 12
   3566: 'Spare_Fault_3566', class No Acknowledgement, trigger "DB302_HMI_Faults_Carrier55_Faults_2" bit 13
   3567: 'Spare_Fault_3567', class No Acknowledgement, trigger "DB302_HMI_Faults_Carrier55_Faults_2" bit 14
   3568: 'Spare_Fault_3568', class No Acknowledgement, trigger "DB302_HMI_Faults_Carrier55_Faults_2" bit 15
   3569: 'Spare_Fault_3569', class No Acknowledgement, trigger "DB302_HMI_Faults_Carrier55_Faults_3" bit 0
   3570: 'Spare_Fault_3570', class No Acknowledgement, trigger "DB302_HMI_Faults_Carrier55_Faults_3" bit 1
   3571: 'Spare_Fault_3571', class No Acknowledgement, trigger "DB302_HMI_Faults_Carrier55_Faults_3" bit 2
   3572: 'Spare_Fault_3572', class No Acknowledgement, trigger "DB302_HMI_Faults_Carrier55_Faults_3" bit 3
   3573: 'Spare_Fault_3573', class No Acknowledgement, trigger "DB302_HMI_Faults_Carrier55_Faults_3" bit 4
   3574: 'Spare_Fault_3574', class No Acknowledgement, trigger "DB302_HMI_Faults_Carrier55_Faults_3" bit 5
   3575: 'Spare_Fault_3575', class No Acknowledgement, trigger "DB302_HMI_Faults_Carrier55_Faults_3" bit 6
   3576: 'Spare_Fault_3576', class No Acknowledgement, trigger "DB302_HMI_Faults_Carrier55_Faults_3" bit 7
   3577: 'Spare_Fault_3577', class No Acknowledgement, trigger "DB302_HMI_Faults_Carrier55_Faults_3" bit 8
   3578: 'Spare_Fault_3578', class No Acknowledgement, trigger "DB302_HMI_Faults_Carrier55_Faults_3" bit 9
   3579: 'Spare_Fault_3579', class No Acknowledgement, trigger "DB302_HMI_Faults_Carrier55_Faults_3" bit 10
   3580: 'Spare_Fault_3580', class No Acknowledgement, trigger "DB302_HMI_Faults_Carrier55_Faults_3" bit 11
   3581: 'Spare_Fault_3581', class No Acknowledgement, trigger "DB302_HMI_Faults_Carrier55_Faults_3" bit 12
   3582: 'Spare_Fault_3582', class No Acknowledgement, trigger "DB302_HMI_Faults_Carrier55_Faults_3" bit 13
   3583: 'Spare_Fault_3583', class No Acknowledgement, trigger "DB302_HMI_Faults_Carrier55_Faults_3" bit 14
   3584: 'Spare_Fault_3584', class No Acknowledgement, trigger "DB302_HMI_Faults_Carrier55_Faults_3" bit 15
   3585: 'Carrier 56 Disconnect Open Power Fault DI11.0', class No Acknowledgement, trigger "DB302_HMI_Faults_Carrier56_Faults_0" bit 0
   3586: 'Carrier 56 Drive Profinet Comm Fault', class No Acknowledgement, trigger "DB302_HMI_Faults_Carrier56_Faults_0" bit 1
   3587: 'Carrier 56 Production Stop Not Reset', class No Acknowledgement, trigger "DB302_HMI_Faults_Carrier56_Faults_0" bit 2
   3588: 'Carrier 56 CB02122 Tripped', class No Acknowledgement, trigger "DB302_HMI_Faults_Carrier56_Faults_0" bit 3
   3589: 'Carrier 56 CB02123 Tripped', class No Acknowledgement, trigger "DB302_HMI_Faults_Carrier56_Faults_0" bit 4
   3590: 'Carrier 56 AUX1 CB Tripped', class No Acknowledgement, trigger "DB302_HMI_Faults_Carrier56_Faults_0" bit 5
   3591: 'Carrier 56 AUX2 CB Tripped', class No Acknowledgement, trigger "DB302_HMI_Faults_Carrier56_Faults_0" bit 6
   3592: 'Carrier 56 PLC Not Communicating', class No Acknowledgement, trigger "DB302_HMI_Faults_Carrier56_Faults_0" bit 7
   3593: 'Carrier 56 Safe Input Card Fault', class No Acknowledgement, trigger "DB302_HMI_Faults_Carrier56_Faults_0" bit 8
   3594: 'Carrier 56 Safe Output Card Fault', class No Acknowledgement, trigger "DB302_HMI_Faults_Carrier56_Faults_0" bit 9
   3595: 'Carrier 56 Standard Input Card Fault', class No Acknowledgement, trigger "DB302_HMI_Faults_Carrier56_Faults_0" bit 10
   3596: 'Carrier 56 Standard Output Card Fault', class No Acknowledgement, trigger "DB302_HMI_Faults_Carrier56_Faults_0" bit 11
   3597: 'Carrier 56 Encoder Position Fault', class No Acknowledgement, trigger "DB302_HMI_Faults_Carrier56_Faults_0" bit 12
   3598: 'Carrier 56 Encoder Internal Error', class No Acknowledgement, trigger "DB302_HMI_Faults_Carrier56_Faults_0" bit 13
   3599: 'Carrier 56 Encoder Comm Fault', class No Acknowledgement, trigger "DB302_HMI_Faults_Carrier56_Faults_0" bit 14
   3600: 'Carrier 56 HMI Comm Fault', class No Acknowledgement, trigger "DB302_HMI_Faults_Carrier56_Faults_0" bit 15
   3601: 'Carrier 56 Crash Detection Fault', class No Acknowledgement, trigger "DB302_HMI_Faults_Carrier56_Faults_1" bit 0
   3602: 'Carrier 56 Carrier Number Invalid', class No Acknowledgement, trigger "DB302_HMI_Faults_Carrier56_Faults_1" bit 1
   3603: 'Carrier 56 Drive: PROFINET configuration error', class No Acknowledgement, trigger "DB302_HMI_Faults_Carrier56_Faults_1" bit 2
   3604: 'Carrier 56 Drive: Error internal communications', class No Acknowledgement, trigger "DB302_HMI_Faults_Carrier56_Faults_1" bit 3
   3605: 'Carrier 56 Drive: Motor overtemperature', class No Acknowledgement, trigger "DB302_HMI_Faults_Carrier56_Faults_1" bit 4
   3606: 'Carrier 56 Drive: Motor overcurrent', class No Acknowledgement, trigger "DB302_HMI_Faults_Carrier56_Faults_1" bit 5
   3607: 'Carrier 56 Drive: Infeed or power unit not ready', class No Acknowledgement, trigger "DB302_HMI_Faults_Carrier56_Faults_1" bit 6
   3608: 'Carrier 56 Drive: Short-circuit/ground fault detected', class No Acknowledgement, trigger "DB302_HMI_Faults_Carrier56_Faults_1" bit 7
   3609: 'Carrier 56 Drive: PROFINET Setpoint timeout', class No Acknowledgement, trigger "DB302_HMI_Faults_Carrier56_Faults_1" bit 8
   3610: 'Carrier 56 Power unit: Overcurrent', class No Acknowledgement, trigger "DB302_HMI_Faults_Carrier56_Faults_1" bit 9
   3611: 'Carrier 56 Power unit: DC link voltage overvoltage', class No Acknowledgement, trigger "DB302_HMI_Faults_Carrier56_Faults_1" bit 10
   3612: 'Carrier 56 Power unit: DC link voltage undervoltage', class No Acknowledgement, trigger "DB302_HMI_Faults_Carrier56_Faults_1" bit 11
   3613: 'Carrier 56 Power unit: Line phase failure in main circuit', class No Acknowledgement, trigger "DB302_HMI_Faults_Carrier56_Faults_1" bit 12
   3614: 'Carrier 56 Power unit: Phase failure motor cable', class No Acknowledgement, trigger "DB302_HMI_Faults_Carrier56_Faults_1" bit 13
   3615: 'Carrier 56 Power unit: Ground fault', class No Acknowledgement, trigger "DB302_HMI_Faults_Carrier56_Faults_1" bit 14
   3616: 'Spare_Fault_3616', class No Acknowledgement, trigger "DB302_HMI_Faults_Carrier56_Faults_1" bit 15
   3617: 'Carrier 56 Motion Off Fault', class No Acknowledgement, trigger "DB302_HMI_Faults_Carrier56_Faults_2" bit 0
   3618: 'Carrier 56 Motion On Fault', class No Acknowledgement, trigger "DB302_HMI_Faults_Carrier56_Faults_2" bit 1
   3619: 'Carrier 56 Spacing Fault', class No Acknowledgement, trigger "DB302_HMI_Faults_Carrier56_Faults_2" bit 2
   3620: 'Carrier 56 Duplicate Carrier Number Fault', class No Acknowledgement, trigger "DB302_HMI_Faults_Carrier56_Faults_2" bit 3
   3621: 'Spare_Fault_3621', class No Acknowledgement, trigger "DB302_HMI_Faults_Carrier56_Faults_2" bit 4
   3622: 'Spare_Fault_3622', class No Acknowledgement, trigger "DB302_HMI_Faults_Carrier56_Faults_2" bit 5
   3623: 'Spare_Fault_3623', class No Acknowledgement, trigger "DB302_HMI_Faults_Carrier56_Faults_2" bit 6
   3624: 'Spare_Fault_3624', class No Acknowledgement, trigger "DB302_HMI_Faults_Carrier56_Faults_2" bit 7
   3625: 'Spare_Fault_3625', class No Acknowledgement, trigger "DB302_HMI_Faults_Carrier56_Faults_2" bit 8
   3626: 'Spare_Fault_3626', class No Acknowledgement, trigger "DB302_HMI_Faults_Carrier56_Faults_2" bit 9
   3627: 'Spare_Fault_3627', class No Acknowledgement, trigger "DB302_HMI_Faults_Carrier56_Faults_2" bit 10
   3628: 'Spare_Fault_3628', class No Acknowledgement, trigger "DB302_HMI_Faults_Carrier56_Faults_2" bit 11
   3629: 'Spare_Fault_3629', class No Acknowledgement, trigger "DB302_HMI_Faults_Carrier56_Faults_2" bit 12
   3630: 'Spare_Fault_3630', class No Acknowledgement, trigger "DB302_HMI_Faults_Carrier56_Faults_2" bit 13
   3631: 'Spare_Fault_3631', class No Acknowledgement, trigger "DB302_HMI_Faults_Carrier56_Faults_2" bit 14
   3632: 'Spare_Fault_3632', class No Acknowledgement, trigger "DB302_HMI_Faults_Carrier56_Faults_2" bit 15
   3633: 'Spare_Fault_3633', class No Acknowledgement, trigger "DB302_HMI_Faults_Carrier56_Faults_3" bit 0
   3634: 'Spare_Fault_3634', class No Acknowledgement, trigger "DB302_HMI_Faults_Carrier56_Faults_3" bit 1
   3635: 'Spare_Fault_3635', class No Acknowledgement, trigger "DB302_HMI_Faults_Carrier56_Faults_3" bit 2
   3636: 'Spare_Fault_3636', class No Acknowledgement, trigger "DB302_HMI_Faults_Carrier56_Faults_3" bit 3
   3637: 'Spare_Fault_3637', class No Acknowledgement, trigger "DB302_HMI_Faults_Carrier56_Faults_3" bit 4
   3638: 'Spare_Fault_3638', class No Acknowledgement, trigger "DB302_HMI_Faults_Carrier56_Faults_3" bit 5
   3639: 'Spare_Fault_3639', class No Acknowledgement, trigger "DB302_HMI_Faults_Carrier56_Faults_3" bit 6
   3640: 'Spare_Fault_3640', class No Acknowledgement, trigger "DB302_HMI_Faults_Carrier56_Faults_3" bit 7
   3641: 'Spare_Fault_3641', class No Acknowledgement, trigger "DB302_HMI_Faults_Carrier56_Faults_3" bit 8
   3642: 'Spare_Fault_3642', class No Acknowledgement, trigger "DB302_HMI_Faults_Carrier56_Faults_3" bit 9
   3643: 'Spare_Fault_3643', class No Acknowledgement, trigger "DB302_HMI_Faults_Carrier56_Faults_3" bit 10
   3644: 'Spare_Fault_3644', class No Acknowledgement, trigger "DB302_HMI_Faults_Carrier56_Faults_3" bit 11
   3645: 'Spare_Fault_3645', class No Acknowledgement, trigger "DB302_HMI_Faults_Carrier56_Faults_3" bit 12
   3646: 'Spare_Fault_3646', class No Acknowledgement, trigger "DB302_HMI_Faults_Carrier56_Faults_3" bit 13
   3647: 'Spare_Fault_3647', class No Acknowledgement, trigger "DB302_HMI_Faults_Carrier56_Faults_3" bit 14